REGION Network 126: DB2062.DBX17.2/3 = LT422 1P Tank Level
   // BTCS_ALARM_WORD_09_BIT_10/11                      14.13
   RUNG wire#powerrail
      "LT422 1P  TANK LEVEL ALARM"(Enable := wire#w1, Value := "20_TANKS_IP_DATA".RIO_01.SECOND_TANK.BWT_LEVEL, "Raw Value" := "IN_Level_WBT_1P", "Enable Delay Time" := "2086_Times"."Alarm Enable Delay", "High Value Release" := false, "SHORT CIRCUIT VALUE" :=, "BROKEN WIRE VALUE" :=, "VERY LOW LEVEL VALUE (LL)" :=, "LOW LEVEL VALUE (L)" := "2084_Setpoints".LT422_Lo, "HIGH LEVEL VALUE (H)" := "2084_Setpoints".LT422_Hi, "VERY HIGH LEVEL VALUE (HH)" := 32000.0, OFFSET :=, "ALARM DELAY" := "2086_Times"."LT422 Alarm Delay", "Peak Value Reset" :=, "ALARM HH" =>, "ALARM H" =>, "ALARM L" =>, "ALARM LL" =>, "ALARM READING" => %DB2062.DBX367.5, "Peak Value" =>, Alarm =>, Alarm_INT =>)   // Raw value not available for Out of Range determination
      wire#w2
      Contact( "LT422 1P  TANK LEVEL ALARM"."ALARM H" )
      Coil( %DB2062.DBX17.2 )
   END_RUNG
   RUNG wire#powerrail
      I_Contact( "2062_Warning_Data"."Water Level Override 1P" )
      { S7_Templates := "SrcType := Int" } GT_Contact(in1 := "504_Tank Grouping_DB2020"."GROUP of TANK 2", in2 := 0)
   END_RUNG wire#w1
   RUNG wire#w2
      Contact( "LT422 1P  TANK LEVEL ALARM"."ALARM L" )
      Coil( %DB2062.DBX17.3 )
   END_RUNG
   // the same network as SCL:
   "LT422 1P  TANK LEVEL ALARM"(Value := "20_TANKS_IP_DATA".RIO_01.SECOND_TANK.BWT_LEVEL,   // "502_ALM_ANALOG": Raw value not available for Out of Range determination
                           "Raw Value" := "IN_Level_WBT_1P",
                           Enable := NOT "2062_Warning_Data"."Water Level Override 1P" AND ("504_Tank Grouping_DB2020"."GROUP of TANK 2" > 0),
                           "Enable Delay Time" := "2086_Times"."Alarm Enable Delay",
                           "High Value Release" := false,
                           "LOW LEVEL VALUE (L)" := "2084_Setpoints".LT422_Lo,
                           "HIGH LEVEL VALUE (H)" := "2084_Setpoints".LT422_Hi,
                           "VERY HIGH LEVEL VALUE (HH)" := 32000.0,
                           "ALARM DELAY" := "2086_Times"."LT422 Alarm Delay",
                           "ALARM READING" => %DB2062.DBX367.5,
                           ENO => #_w1);
   %DB2062.DBX17.2 := #_w1 AND "LT422 1P  TANK LEVEL ALARM"."ALARM H";
   %DB2062.DBX17.3 := #_w1 AND "LT422 1P  TANK LEVEL ALARM"."ALARM L";
END_REGION

REGION Network 127: DB2062.DBX17.4/5 = LT421 1S Tank Level
   // BTCS_ALARM_WORD_09_BIT_12/13                                  14.14
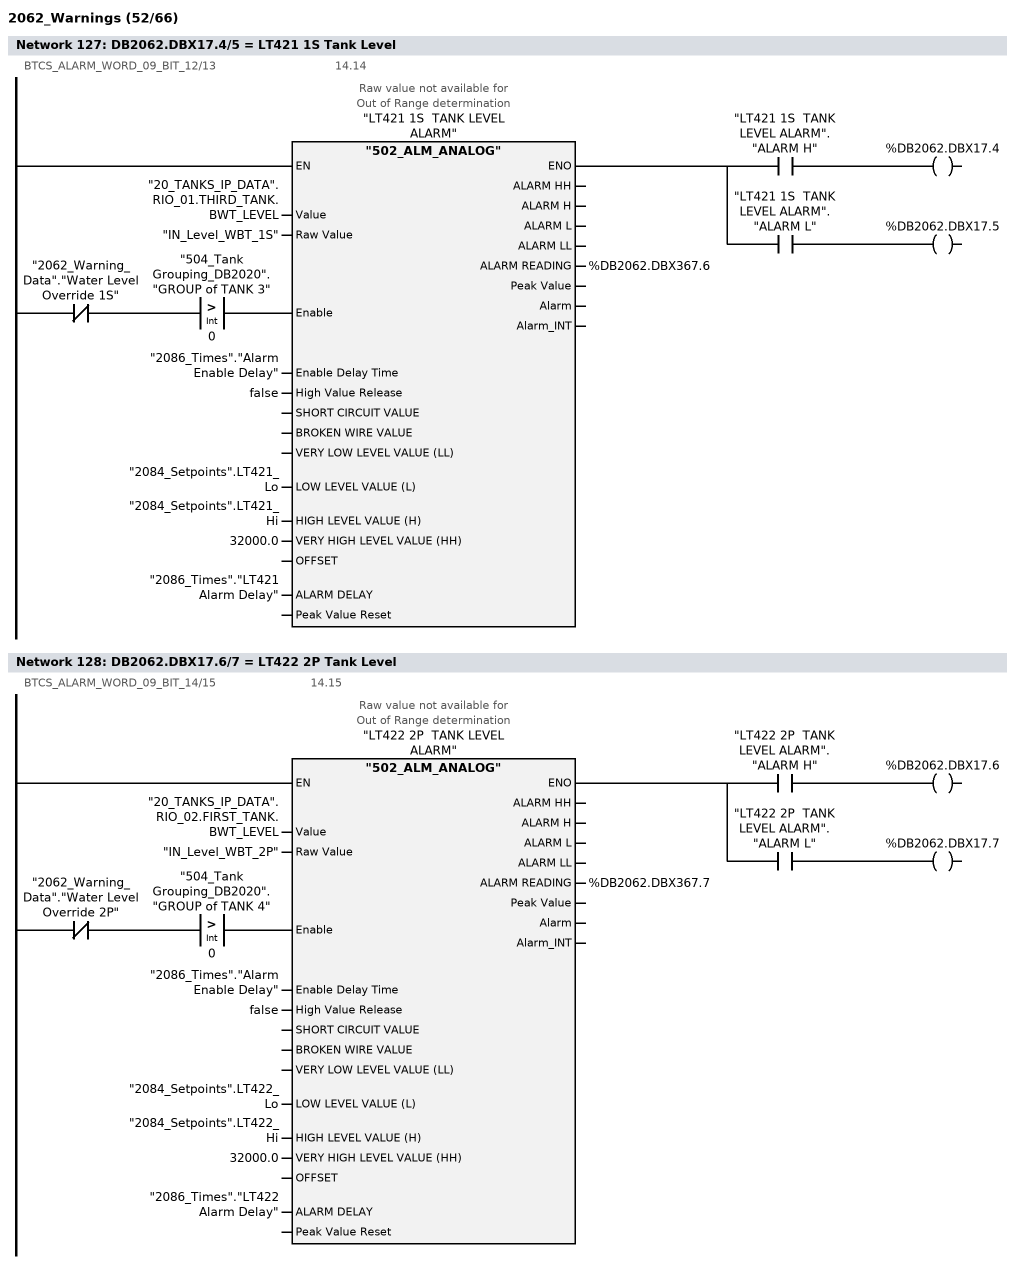
   RUNG wire#powerrail
      "LT421 1S  TANK LEVEL ALARM"(Enable := wire#w1, Value := "20_TANKS_IP_DATA".RIO_01.THIRD_TANK.BWT_LEVEL, "Raw Value" := "IN_Level_WBT_1S", "Enable Delay Time" := "2086_Times"."Alarm Enable Delay", "High Value Release" := false, "SHORT CIRCUIT VALUE" :=, "BROKEN WIRE VALUE" :=, "VERY LOW LEVEL VALUE (LL)" :=, "LOW LEVEL VALUE (L)" := "2084_Setpoints".LT421_Lo, "HIGH LEVEL VALUE (H)" := "2084_Setpoints".LT421_Hi, "VERY HIGH LEVEL VALUE (HH)" := 32000.0, OFFSET :=, "ALARM DELAY" := "2086_Times"."LT421 Alarm Delay", "Peak Value Reset" :=, "ALARM HH" =>, "ALARM H" =>, "ALARM L" =>, "ALARM LL" =>, "ALARM READING" => %DB2062.DBX367.6, "Peak Value" =>, Alarm =>, Alarm_INT =>)   // Raw value not available for Out of Range determination
      wire#w2
      Contact( "LT421 1S  TANK LEVEL ALARM"."ALARM H" )
      Coil( %DB2062.DBX17.4 )
   END_RUNG
   RUNG wire#powerrail
      I_Contact( "2062_Warning_Data"."Water Level Override 1S" )
      { S7_Templates := "SrcType := Int" } GT_Contact(in1 := "504_Tank Grouping_DB2020"."GROUP of TANK 3", in2 := 0)
   END_RUNG wire#w1
   RUNG wire#w2
      Contact( "LT421 1S  TANK LEVEL ALARM"."ALARM L" )
      Coil( %DB2062.DBX17.5 )
   END_RUNG
   // the same network as SCL:
   "LT421 1S  TANK LEVEL ALARM"(Value := "20_TANKS_IP_DATA".RIO_01.THIRD_TANK.BWT_LEVEL,   // "502_ALM_ANALOG": Raw value not available for Out of Range determination
                           "Raw Value" := "IN_Level_WBT_1S",
                           Enable := NOT "2062_Warning_Data"."Water Level Override 1S" AND ("504_Tank Grouping_DB2020"."GROUP of TANK 3" > 0),
                           "Enable Delay Time" := "2086_Times"."Alarm Enable Delay",
                           "High Value Release" := false,
                           "LOW LEVEL VALUE (L)" := "2084_Setpoints".LT421_Lo,
                           "HIGH LEVEL VALUE (H)" := "2084_Setpoints".LT421_Hi,
                           "VERY HIGH LEVEL VALUE (HH)" := 32000.0,
                           "ALARM DELAY" := "2086_Times"."LT421 Alarm Delay",
                           "ALARM READING" => %DB2062.DBX367.6,
                           ENO => #_w1);
   %DB2062.DBX17.4 := #_w1 AND "LT421 1S  TANK LEVEL ALARM"."ALARM H";
   %DB2062.DBX17.5 := #_w1 AND "LT421 1S  TANK LEVEL ALARM"."ALARM L";
END_REGION

REGION Network 128: DB2062.DBX17.6/7 = LT422 2P Tank Level
   // BTCS_ALARM_WORD_09_BIT_14/15                           14.15
   RUNG wire#powerrail
      "LT422 2P  TANK LEVEL ALARM"(Enable := wire#w1, Value := "20_TANKS_IP_DATA".RIO_02.FIRST_TANK.BWT_LEVEL, "Raw Value" := "IN_Level_WBT_2P", "Enable Delay Time" := "2086_Times"."Alarm Enable Delay", "High Value Release" := false, "SHORT CIRCUIT VALUE" :=, "BROKEN WIRE VALUE" :=, "VERY LOW LEVEL VALUE (LL)" :=, "LOW LEVEL VALUE (L)" := "2084_Setpoints".LT422_Lo, "HIGH LEVEL VALUE (H)" := "2084_Setpoints".LT422_Hi, "VERY HIGH LEVEL VALUE (HH)" := 32000.0, OFFSET :=, "ALARM DELAY" := "2086_Times"."LT422 Alarm Delay", "Peak Value Reset" :=, "ALARM HH" =>, "ALARM H" =>, "ALARM L" =>, "ALARM LL" =>, "ALARM READING" => %DB2062.DBX367.7, "Peak Value" =>, Alarm =>, Alarm_INT =>)   // Raw value not available for Out of Range determination
      wire#w2
      Contact( "LT422 2P  TANK LEVEL ALARM"."ALARM H" )
      Coil( %DB2062.DBX17.6 )
   END_RUNG
   RUNG wire#powerrail
      I_Contact( "2062_Warning_Data"."Water Level Override 2P" )
      { S7_Templates := "SrcType := Int" } GT_Contact(in1 := "504_Tank Grouping_DB2020"."GROUP of TANK 4", in2 := 0)
   END_RUNG wire#w1
   RUNG wire#w2
      Contact( "LT422 2P  TANK LEVEL ALARM"."ALARM L" )
      Coil( %DB2062.DBX17.7 )
   END_RUNG
   // the same network as SCL:
   "LT422 2P  TANK LEVEL ALARM"(Value := "20_TANKS_IP_DATA".RIO_02.FIRST_TANK.BWT_LEVEL,   // "502_ALM_ANALOG": Raw value not available for Out of Range determination
                           "Raw Value" := "IN_Level_WBT_2P",
                           Enable := NOT "2062_Warning_Data"."Water Level Override 2P" AND ("504_Tank Grouping_DB2020"."GROUP of TANK 4" > 0),
                           "Enable Delay Time" := "2086_Times"."Alarm Enable Delay",
                           "High Value Release" := false,
                           "LOW LEVEL VALUE (L)" := "2084_Setpoints".LT422_Lo,
                           "HIGH LEVEL VALUE (H)" := "2084_Setpoints".LT422_Hi,
                           "VERY HIGH LEVEL VALUE (HH)" := 32000.0,
                           "ALARM DELAY" := "2086_Times"."LT422 Alarm Delay",
                           "ALARM READING" => %DB2062.DBX367.7,
                           ENO => #_w1);
   %DB2062.DBX17.6 := #_w1 AND "LT422 2P  TANK LEVEL ALARM"."ALARM H";
   %DB2062.DBX17.7 := #_w1 AND "LT422 2P  TANK LEVEL ALARM"."ALARM L";
END_REGION

REGION Network 129: DB2062.DBX18.0/1 = LT421 2S Tank Level
   // BTCS_ALARM_WORD_10_BIT_0/1                                    15.0
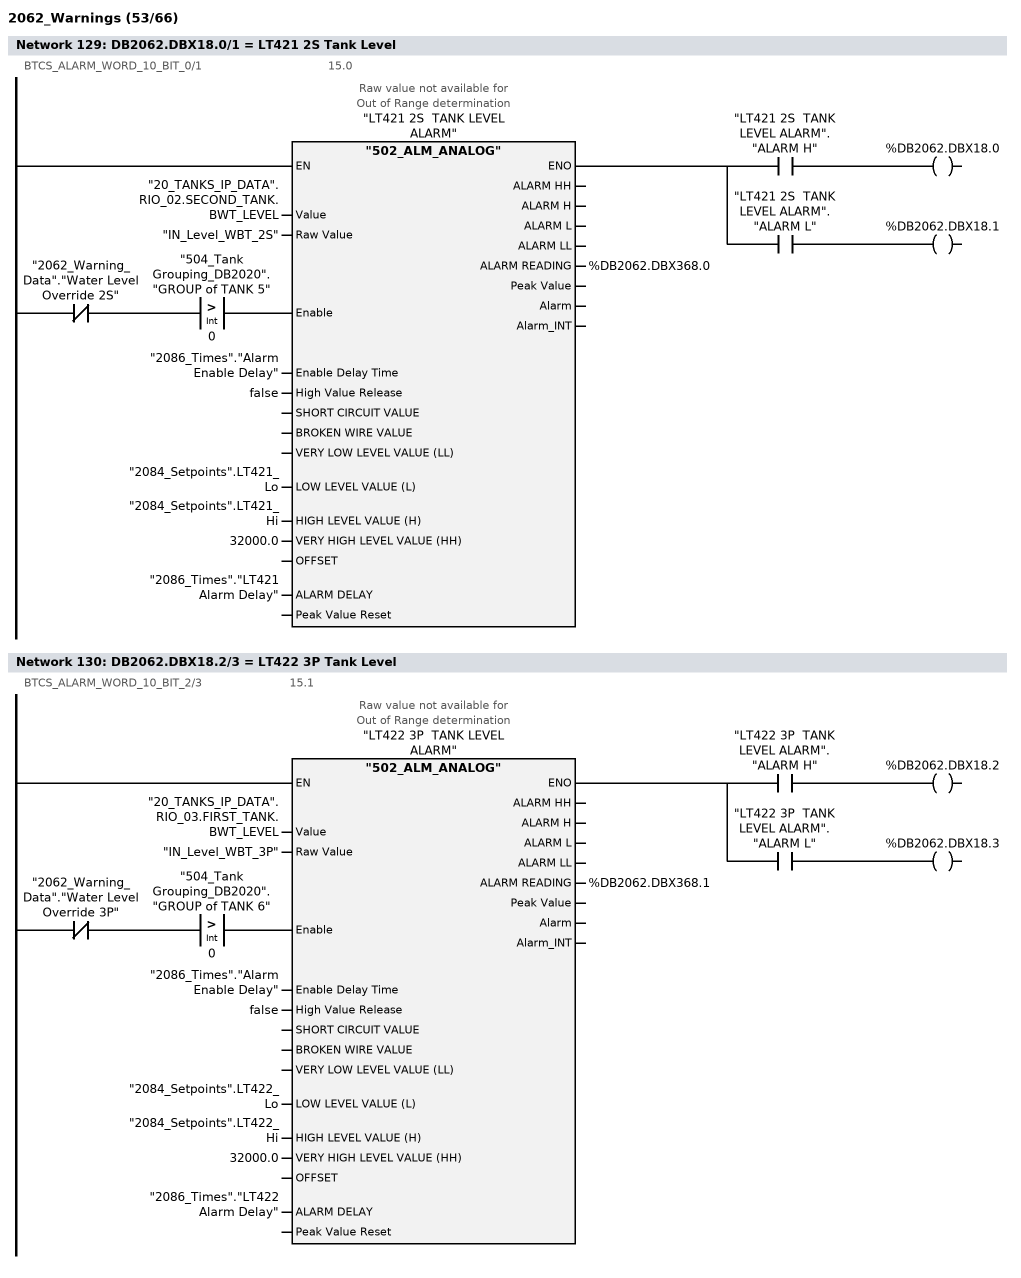
   RUNG wire#powerrail
      "LT421 2S  TANK LEVEL ALARM"(Enable := wire#w1, Value := "20_TANKS_IP_DATA".RIO_02.SECOND_TANK.BWT_LEVEL, "Raw Value" := "IN_Level_WBT_2S", "Enable Delay Time" := "2086_Times"."Alarm Enable Delay", "High Value Release" := false, "SHORT CIRCUIT VALUE" :=, "BROKEN WIRE VALUE" :=, "VERY LOW LEVEL VALUE (LL)" :=, "LOW LEVEL VALUE (L)" := "2084_Setpoints".LT421_Lo, "HIGH LEVEL VALUE (H)" := "2084_Setpoints".LT421_Hi, "VERY HIGH LEVEL VALUE (HH)" := 32000.0, OFFSET :=, "ALARM DELAY" := "2086_Times"."LT421 Alarm Delay", "Peak Value Reset" :=, "ALARM HH" =>, "ALARM H" =>, "ALARM L" =>, "ALARM LL" =>, "ALARM READING" => %DB2062.DBX368.0, "Peak Value" =>, Alarm =>, Alarm_INT =>)   // Raw value not available for Out of Range determination
      wire#w2
      Contact( "LT421 2S  TANK LEVEL ALARM"."ALARM H" )
      Coil( %DB2062.DBX18.0 )
   END_RUNG
   RUNG wire#powerrail
      I_Contact( "2062_Warning_Data"."Water Level Override 2S" )
      { S7_Templates := "SrcType := Int" } GT_Contact(in1 := "504_Tank Grouping_DB2020"."GROUP of TANK 5", in2 := 0)
   END_RUNG wire#w1
   RUNG wire#w2
      Contact( "LT421 2S  TANK LEVEL ALARM"."ALARM L" )
      Coil( %DB2062.DBX18.1 )
   END_RUNG
   // the same network as SCL:
   "LT421 2S  TANK LEVEL ALARM"(Value := "20_TANKS_IP_DATA".RIO_02.SECOND_TANK.BWT_LEVEL,   // "502_ALM_ANALOG": Raw value not available for Out of Range determination
                           "Raw Value" := "IN_Level_WBT_2S",
                           Enable := NOT "2062_Warning_Data"."Water Level Override 2S" AND ("504_Tank Grouping_DB2020"."GROUP of TANK 5" > 0),
                           "Enable Delay Time" := "2086_Times"."Alarm Enable Delay",
                           "High Value Release" := false,
                           "LOW LEVEL VALUE (L)" := "2084_Setpoints".LT421_Lo,
                           "HIGH LEVEL VALUE (H)" := "2084_Setpoints".LT421_Hi,
                           "VERY HIGH LEVEL VALUE (HH)" := 32000.0,
                           "ALARM DELAY" := "2086_Times"."LT421 Alarm Delay",
                           "ALARM READING" => %DB2062.DBX368.0,
                           ENO => #_w1);
   %DB2062.DBX18.0 := #_w1 AND "LT421 2S  TANK LEVEL ALARM"."ALARM H";
   %DB2062.DBX18.1 := #_w1 AND "LT421 2S  TANK LEVEL ALARM"."ALARM L";
END_REGION

REGION Network 130: DB2062.DBX18.2/3 = LT422 3P Tank Level
   // BTCS_ALARM_WORD_10_BIT_2/3                         15.1
   RUNG wire#powerrail
      "LT422 3P  TANK LEVEL ALARM"(Enable := wire#w1, Value := "20_TANKS_IP_DATA".RIO_03.FIRST_TANK.BWT_LEVEL, "Raw Value" := "IN_Level_WBT_3P", "Enable Delay Time" := "2086_Times"."Alarm Enable Delay", "High Value Release" := false, "SHORT CIRCUIT VALUE" :=, "BROKEN WIRE VALUE" :=, "VERY LOW LEVEL VALUE (LL)" :=, "LOW LEVEL VALUE (L)" := "2084_Setpoints".LT422_Lo, "HIGH LEVEL VALUE (H)" := "2084_Setpoints".LT422_Hi, "VERY HIGH LEVEL VALUE (HH)" := 32000.0, OFFSET :=, "ALARM DELAY" := "2086_Times"."LT422 Alarm Delay", "Peak Value Reset" :=, "ALARM HH" =>, "ALARM H" =>, "ALARM L" =>, "ALARM LL" =>, "ALARM READING" => %DB2062.DBX368.1, "Peak Value" =>, Alarm =>, Alarm_INT =>)   // Raw value not available for Out of Range determination
      wire#w2
      Contact( "LT422 3P  TANK LEVEL ALARM"."ALARM H" )
      Coil( %DB2062.DBX18.2 )
   END_RUNG
   RUNG wire#powerrail
      I_Contact( "2062_Warning_Data"."Water Level Override 3P" )
      { S7_Templates := "SrcType := Int" } GT_Contact(in1 := "504_Tank Grouping_DB2020"."GROUP of TANK 6", in2 := 0)
   END_RUNG wire#w1
   RUNG wire#w2
      Contact( "LT422 3P  TANK LEVEL ALARM"."ALARM L" )
      Coil( %DB2062.DBX18.3 )
   END_RUNG
   // the same network as SCL:
   "LT422 3P  TANK LEVEL ALARM"(Value := "20_TANKS_IP_DATA".RIO_03.FIRST_TANK.BWT_LEVEL,   // "502_ALM_ANALOG": Raw value not available for Out of Range determination
                           "Raw Value" := "IN_Level_WBT_3P",
                           Enable := NOT "2062_Warning_Data"."Water Level Override 3P" AND ("504_Tank Grouping_DB2020"."GROUP of TANK 6" > 0),
                           "Enable Delay Time" := "2086_Times"."Alarm Enable Delay",
                           "High Value Release" := false,
                           "LOW LEVEL VALUE (L)" := "2084_Setpoints".LT422_Lo,
                           "HIGH LEVEL VALUE (H)" := "2084_Setpoints".LT422_Hi,
                           "VERY HIGH LEVEL VALUE (HH)" := 32000.0,
                           "ALARM DELAY" := "2086_Times"."LT422 Alarm Delay",
                           "ALARM READING" => %DB2062.DBX368.1,
                           ENO => #_w1);
   %DB2062.DBX18.2 := #_w1 AND "LT422 3P  TANK LEVEL ALARM"."ALARM H";
   %DB2062.DBX18.3 := #_w1 AND "LT422 3P  TANK LEVEL ALARM"."ALARM L";
END_REGION

REGION Network 131: DB2062.DBX18.4/5 = LT421 3S Tank Level
   // BTCS_ALARM_WORD_10_BIT_4/5                               15.2
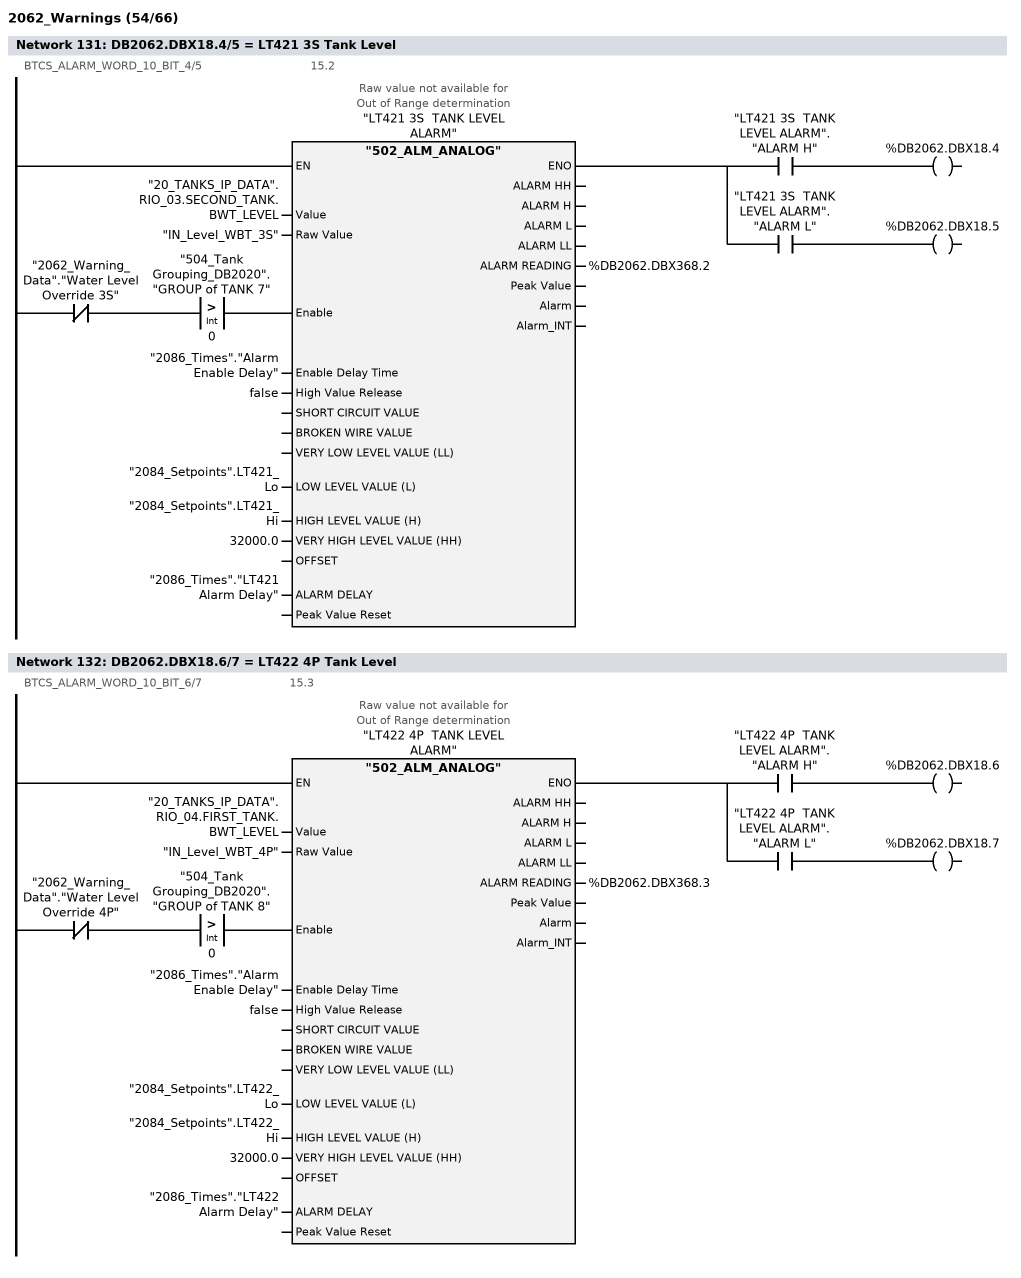
   RUNG wire#powerrail
      "LT421 3S  TANK LEVEL ALARM"(Enable := wire#w1, Value := "20_TANKS_IP_DATA".RIO_03.SECOND_TANK.BWT_LEVEL, "Raw Value" := "IN_Level_WBT_3S", "Enable Delay Time" := "2086_Times"."Alarm Enable Delay", "High Value Release" := false, "SHORT CIRCUIT VALUE" :=, "BROKEN WIRE VALUE" :=, "VERY LOW LEVEL VALUE (LL)" :=, "LOW LEVEL VALUE (L)" := "2084_Setpoints".LT421_Lo, "HIGH LEVEL VALUE (H)" := "2084_Setpoints".LT421_Hi, "VERY HIGH LEVEL VALUE (HH)" := 32000.0, OFFSET :=, "ALARM DELAY" := "2086_Times"."LT421 Alarm Delay", "Peak Value Reset" :=, "ALARM HH" =>, "ALARM H" =>, "ALARM L" =>, "ALARM LL" =>, "ALARM READING" => %DB2062.DBX368.2, "Peak Value" =>, Alarm =>, Alarm_INT =>)   // Raw value not available for Out of Range determination
      wire#w2
      Contact( "LT421 3S  TANK LEVEL ALARM"."ALARM H" )
      Coil( %DB2062.DBX18.4 )
   END_RUNG
   RUNG wire#powerrail
      I_Contact( "2062_Warning_Data"."Water Level Override 3S" )
      { S7_Templates := "SrcType := Int" } GT_Contact(in1 := "504_Tank Grouping_DB2020"."GROUP of TANK 7", in2 := 0)
   END_RUNG wire#w1
   RUNG wire#w2
      Contact( "LT421 3S  TANK LEVEL ALARM"."ALARM L" )
      Coil( %DB2062.DBX18.5 )
   END_RUNG
   // the same network as SCL:
   "LT421 3S  TANK LEVEL ALARM"(Value := "20_TANKS_IP_DATA".RIO_03.SECOND_TANK.BWT_LEVEL,   // "502_ALM_ANALOG": Raw value not available for Out of Range determination
                           "Raw Value" := "IN_Level_WBT_3S",
                           Enable := NOT "2062_Warning_Data"."Water Level Override 3S" AND ("504_Tank Grouping_DB2020"."GROUP of TANK 7" > 0),
                           "Enable Delay Time" := "2086_Times"."Alarm Enable Delay",
                           "High Value Release" := false,
                           "LOW LEVEL VALUE (L)" := "2084_Setpoints".LT421_Lo,
                           "HIGH LEVEL VALUE (H)" := "2084_Setpoints".LT421_Hi,
                           "VERY HIGH LEVEL VALUE (HH)" := 32000.0,
                           "ALARM DELAY" := "2086_Times"."LT421 Alarm Delay",
                           "ALARM READING" => %DB2062.DBX368.2,
                           ENO => #_w1);
   %DB2062.DBX18.4 := #_w1 AND "LT421 3S  TANK LEVEL ALARM"."ALARM H";
   %DB2062.DBX18.5 := #_w1 AND "LT421 3S  TANK LEVEL ALARM"."ALARM L";
END_REGION

REGION Network 132: DB2062.DBX18.6/7 = LT422 4P Tank Level
   // BTCS_ALARM_WORD_10_BIT_6/7                         15.3
   RUNG wire#powerrail
      "LT422 4P  TANK LEVEL ALARM"(Enable := wire#w1, Value := "20_TANKS_IP_DATA".RIO_04.FIRST_TANK.BWT_LEVEL, "Raw Value" := "IN_Level_WBT_4P", "Enable Delay Time" := "2086_Times"."Alarm Enable Delay", "High Value Release" := false, "SHORT CIRCUIT VALUE" :=, "BROKEN WIRE VALUE" :=, "VERY LOW LEVEL VALUE (LL)" :=, "LOW LEVEL VALUE (L)" := "2084_Setpoints".LT422_Lo, "HIGH LEVEL VALUE (H)" := "2084_Setpoints".LT422_Hi, "VERY HIGH LEVEL VALUE (HH)" := 32000.0, OFFSET :=, "ALARM DELAY" := "2086_Times"."LT422 Alarm Delay", "Peak Value Reset" :=, "ALARM HH" =>, "ALARM H" =>, "ALARM L" =>, "ALARM LL" =>, "ALARM READING" => %DB2062.DBX368.3, "Peak Value" =>, Alarm =>, Alarm_INT =>)   // Raw value not available for Out of Range determination
      wire#w2
      Contact( "LT422 4P  TANK LEVEL ALARM"."ALARM H" )
      Coil( %DB2062.DBX18.6 )
   END_RUNG
   RUNG wire#powerrail
      I_Contact( "2062_Warning_Data"."Water Level Override 4P" )
      { S7_Templates := "SrcType := Int" } GT_Contact(in1 := "504_Tank Grouping_DB2020"."GROUP of TANK 8", in2 := 0)
   END_RUNG wire#w1
   RUNG wire#w2
      Contact( "LT422 4P  TANK LEVEL ALARM"."ALARM L" )
      Coil( %DB2062.DBX18.7 )
   END_RUNG
   // the same network as SCL:
   "LT422 4P  TANK LEVEL ALARM"(Value := "20_TANKS_IP_DATA".RIO_04.FIRST_TANK.BWT_LEVEL,   // "502_ALM_ANALOG": Raw value not available for Out of Range determination
                           "Raw Value" := "IN_Level_WBT_4P",
                           Enable := NOT "2062_Warning_Data"."Water Level Override 4P" AND ("504_Tank Grouping_DB2020"."GROUP of TANK 8" > 0),
                           "Enable Delay Time" := "2086_Times"."Alarm Enable Delay",
                           "High Value Release" := false,
                           "LOW LEVEL VALUE (L)" := "2084_Setpoints".LT422_Lo,
                           "HIGH LEVEL VALUE (H)" := "2084_Setpoints".LT422_Hi,
                           "VERY HIGH LEVEL VALUE (HH)" := 32000.0,
                           "ALARM DELAY" := "2086_Times"."LT422 Alarm Delay",
                           "ALARM READING" => %DB2062.DBX368.3,
                           ENO => #_w1);
   %DB2062.DBX18.6 := #_w1 AND "LT422 4P  TANK LEVEL ALARM"."ALARM H";
   %DB2062.DBX18.7 := #_w1 AND "LT422 4P  TANK LEVEL ALARM"."ALARM L";
END_REGION

REGION Network 133: DB2062.DBX19.0/1 = LT421 4S Tank Level
   // BTCS_ALARM_WORD_10_BIT_8/9                     15.4
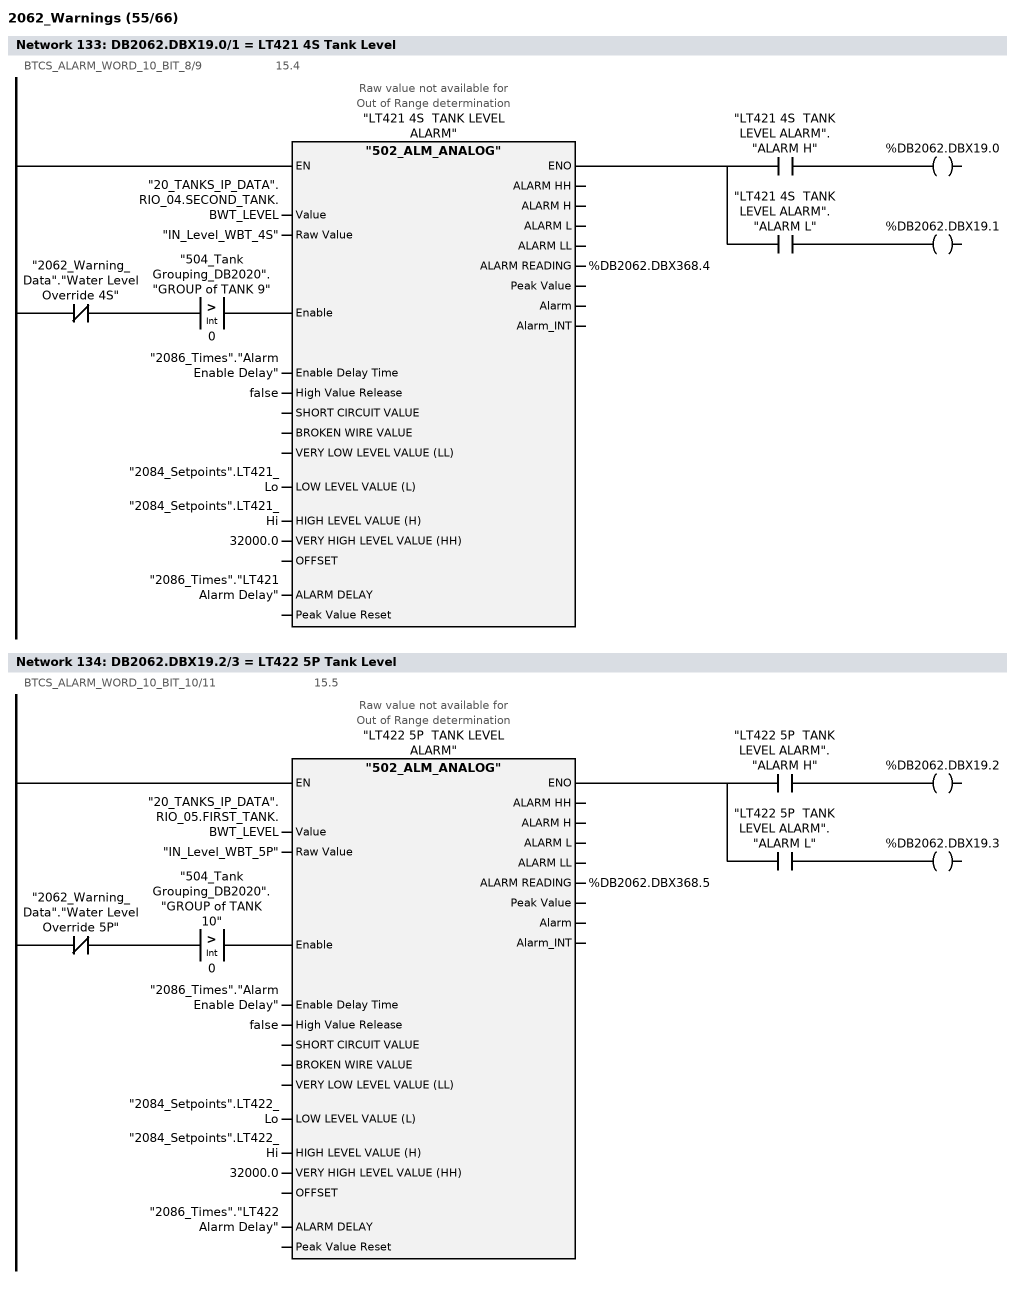
   RUNG wire#powerrail
      "LT421 4S  TANK LEVEL ALARM"(Enable := wire#w1, Value := "20_TANKS_IP_DATA".RIO_04.SECOND_TANK.BWT_LEVEL, "Raw Value" := "IN_Level_WBT_4S", "Enable Delay Time" := "2086_Times"."Alarm Enable Delay", "High Value Release" := false, "SHORT CIRCUIT VALUE" :=, "BROKEN WIRE VALUE" :=, "VERY LOW LEVEL VALUE (LL)" :=, "LOW LEVEL VALUE (L)" := "2084_Setpoints".LT421_Lo, "HIGH LEVEL VALUE (H)" := "2084_Setpoints".LT421_Hi, "VERY HIGH LEVEL VALUE (HH)" := 32000.0, OFFSET :=, "ALARM DELAY" := "2086_Times"."LT421 Alarm Delay", "Peak Value Reset" :=, "ALARM HH" =>, "ALARM H" =>, "ALARM L" =>, "ALARM LL" =>, "ALARM READING" => %DB2062.DBX368.4, "Peak Value" =>, Alarm =>, Alarm_INT =>)   // Raw value not available for Out of Range determination
      wire#w2
      Contact( "LT421 4S  TANK LEVEL ALARM"."ALARM H" )
      Coil( %DB2062.DBX19.0 )
   END_RUNG
   RUNG wire#powerrail
      I_Contact( "2062_Warning_Data"."Water Level Override 4S" )
      { S7_Templates := "SrcType := Int" } GT_Contact(in1 := "504_Tank Grouping_DB2020"."GROUP of TANK 9", in2 := 0)
   END_RUNG wire#w1
   RUNG wire#w2
      Contact( "LT421 4S  TANK LEVEL ALARM"."ALARM L" )
      Coil( %DB2062.DBX19.1 )
   END_RUNG
   // the same network as SCL:
   "LT421 4S  TANK LEVEL ALARM"(Value := "20_TANKS_IP_DATA".RIO_04.SECOND_TANK.BWT_LEVEL,   // "502_ALM_ANALOG": Raw value not available for Out of Range determination
                           "Raw Value" := "IN_Level_WBT_4S",
                           Enable := NOT "2062_Warning_Data"."Water Level Override 4S" AND ("504_Tank Grouping_DB2020"."GROUP of TANK 9" > 0),
                           "Enable Delay Time" := "2086_Times"."Alarm Enable Delay",
                           "High Value Release" := false,
                           "LOW LEVEL VALUE (L)" := "2084_Setpoints".LT421_Lo,
                           "HIGH LEVEL VALUE (H)" := "2084_Setpoints".LT421_Hi,
                           "VERY HIGH LEVEL VALUE (HH)" := 32000.0,
                           "ALARM DELAY" := "2086_Times"."LT421 Alarm Delay",
                           "ALARM READING" => %DB2062.DBX368.4,
                           ENO => #_w1);
   %DB2062.DBX19.0 := #_w1 AND "LT421 4S  TANK LEVEL ALARM"."ALARM H";
   %DB2062.DBX19.1 := #_w1 AND "LT421 4S  TANK LEVEL ALARM"."ALARM L";
END_REGION

REGION Network 134: DB2062.DBX19.2/3 = LT422 5P Tank Level
   // BTCS_ALARM_WORD_10_BIT_10/11                            15.5
   RUNG wire#powerrail
      "LT422 5P  TANK LEVEL ALARM"(Enable := wire#w1, Value := "20_TANKS_IP_DATA".RIO_05.FIRST_TANK.BWT_LEVEL, "Raw Value" := "IN_Level_WBT_5P", "Enable Delay Time" := "2086_Times"."Alarm Enable Delay", "High Value Release" := false, "SHORT CIRCUIT VALUE" :=, "BROKEN WIRE VALUE" :=, "VERY LOW LEVEL VALUE (LL)" :=, "LOW LEVEL VALUE (L)" := "2084_Setpoints".LT422_Lo, "HIGH LEVEL VALUE (H)" := "2084_Setpoints".LT422_Hi, "VERY HIGH LEVEL VALUE (HH)" := 32000.0, OFFSET :=, "ALARM DELAY" := "2086_Times"."LT422 Alarm Delay", "Peak Value Reset" :=, "ALARM HH" =>, "ALARM H" =>, "ALARM L" =>, "ALARM LL" =>, "ALARM READING" => %DB2062.DBX368.5, "Peak Value" =>, Alarm =>, Alarm_INT =>)   // Raw value not available for Out of Range determination
      wire#w2
      Contact( "LT422 5P  TANK LEVEL ALARM"."ALARM H" )
      Coil( %DB2062.DBX19.2 )
   END_RUNG
   RUNG wire#powerrail
      I_Contact( "2062_Warning_Data"."Water Level Override 5P" )
      { S7_Templates := "SrcType := Int" } GT_Contact(in1 := "504_Tank Grouping_DB2020"."GROUP of TANK 10", in2 := 0)
   END_RUNG wire#w1
   RUNG wire#w2
      Contact( "LT422 5P  TANK LEVEL ALARM"."ALARM L" )
      Coil( %DB2062.DBX19.3 )
   END_RUNG
   // the same network as SCL:
   "LT422 5P  TANK LEVEL ALARM"(Value := "20_TANKS_IP_DATA".RIO_05.FIRST_TANK.BWT_LEVEL,   // "502_ALM_ANALOG": Raw value not available for Out of Range determination
                           "Raw Value" := "IN_Level_WBT_5P",
                           Enable := NOT "2062_Warning_Data"."Water Level Override 5P" AND ("504_Tank Grouping_DB2020"."GROUP of TANK 10" > 0),
                           "Enable Delay Time" := "2086_Times"."Alarm Enable Delay",
                           "High Value Release" := false,
                           "LOW LEVEL VALUE (L)" := "2084_Setpoints".LT422_Lo,
                           "HIGH LEVEL VALUE (H)" := "2084_Setpoints".LT422_Hi,
                           "VERY HIGH LEVEL VALUE (HH)" := 32000.0,
                           "ALARM DELAY" := "2086_Times"."LT422 Alarm Delay",
                           "ALARM READING" => %DB2062.DBX368.5,
                           ENO => #_w1);
   %DB2062.DBX19.2 := #_w1 AND "LT422 5P  TANK LEVEL ALARM"."ALARM H";
   %DB2062.DBX19.3 := #_w1 AND "LT422 5P  TANK LEVEL ALARM"."ALARM L";
END_REGION

REGION Network 135: DB2062.DBX19.4/5 = LT421 5S Tank Level
   // BTCS_ALARM_WORD_10_BIT_12/13                          15.6
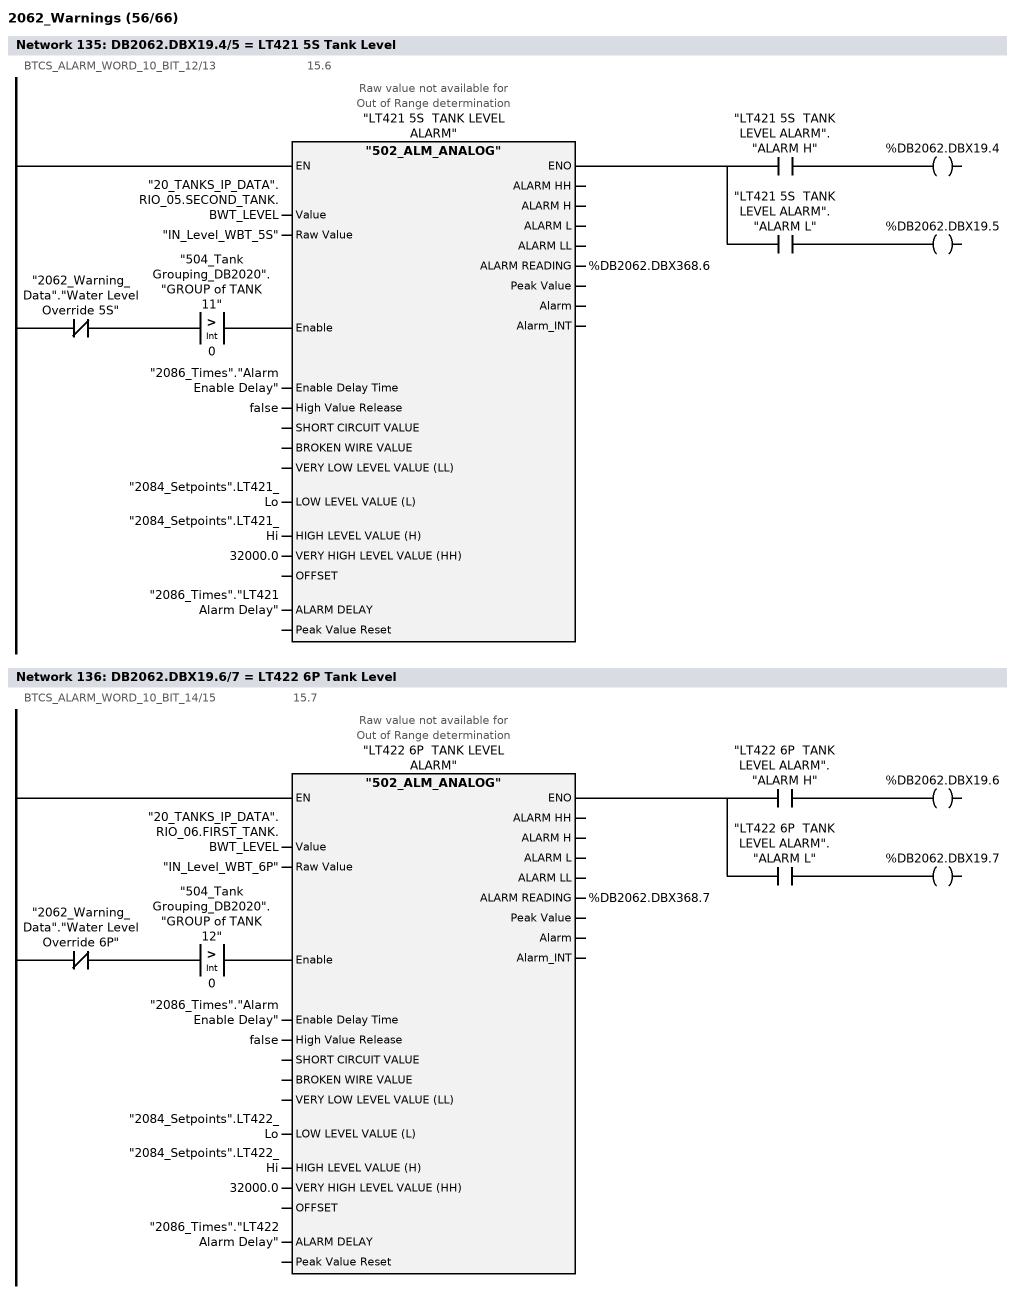
   RUNG wire#powerrail
      "LT421 5S  TANK LEVEL ALARM"(Enable := wire#w1, Value := "20_TANKS_IP_DATA".RIO_05.SECOND_TANK.BWT_LEVEL, "Raw Value" := "IN_Level_WBT_5S", "Enable Delay Time" := "2086_Times"."Alarm Enable Delay", "High Value Release" := false, "SHORT CIRCUIT VALUE" :=, "BROKEN WIRE VALUE" :=, "VERY LOW LEVEL VALUE (LL)" :=, "LOW LEVEL VALUE (L)" := "2084_Setpoints".LT421_Lo, "HIGH LEVEL VALUE (H)" := "2084_Setpoints".LT421_Hi, "VERY HIGH LEVEL VALUE (HH)" := 32000.0, OFFSET :=, "ALARM DELAY" := "2086_Times"."LT421 Alarm Delay", "Peak Value Reset" :=, "ALARM HH" =>, "ALARM H" =>, "ALARM L" =>, "ALARM LL" =>, "ALARM READING" => %DB2062.DBX368.6, "Peak Value" =>, Alarm =>, Alarm_INT =>)   // Raw value not available for Out of Range determination
      wire#w2
      Contact( "LT421 5S  TANK LEVEL ALARM"."ALARM H" )
      Coil( %DB2062.DBX19.4 )
   END_RUNG
   RUNG wire#powerrail
      I_Contact( "2062_Warning_Data"."Water Level Override 5S" )
      { S7_Templates := "SrcType := Int" } GT_Contact(in1 := "504_Tank Grouping_DB2020"."GROUP of TANK 11", in2 := 0)
   END_RUNG wire#w1
   RUNG wire#w2
      Contact( "LT421 5S  TANK LEVEL ALARM"."ALARM L" )
      Coil( %DB2062.DBX19.5 )
   END_RUNG
   // the same network as SCL:
   "LT421 5S  TANK LEVEL ALARM"(Value := "20_TANKS_IP_DATA".RIO_05.SECOND_TANK.BWT_LEVEL,   // "502_ALM_ANALOG": Raw value not available for Out of Range determination
                           "Raw Value" := "IN_Level_WBT_5S",
                           Enable := NOT "2062_Warning_Data"."Water Level Override 5S" AND ("504_Tank Grouping_DB2020"."GROUP of TANK 11" > 0),
                           "Enable Delay Time" := "2086_Times"."Alarm Enable Delay",
                           "High Value Release" := false,
                           "LOW LEVEL VALUE (L)" := "2084_Setpoints".LT421_Lo,
                           "HIGH LEVEL VALUE (H)" := "2084_Setpoints".LT421_Hi,
                           "VERY HIGH LEVEL VALUE (HH)" := 32000.0,
                           "ALARM DELAY" := "2086_Times"."LT421 Alarm Delay",
                           "ALARM READING" => %DB2062.DBX368.6,
                           ENO => #_w1);
   %DB2062.DBX19.4 := #_w1 AND "LT421 5S  TANK LEVEL ALARM"."ALARM H";
   %DB2062.DBX19.5 := #_w1 AND "LT421 5S  TANK LEVEL ALARM"."ALARM L";
END_REGION

REGION Network 136: DB2062.DBX19.6/7 = LT422 6P Tank Level
   // BTCS_ALARM_WORD_10_BIT_14/15                      15.7
   RUNG wire#powerrail
      "LT422 6P  TANK LEVEL ALARM"(Enable := wire#w1, Value := "20_TANKS_IP_DATA".RIO_06.FIRST_TANK.BWT_LEVEL, "Raw Value" := "IN_Level_WBT_6P", "Enable Delay Time" := "2086_Times"."Alarm Enable Delay", "High Value Release" := false, "SHORT CIRCUIT VALUE" :=, "BROKEN WIRE VALUE" :=, "VERY LOW LEVEL VALUE (LL)" :=, "LOW LEVEL VALUE (L)" := "2084_Setpoints".LT422_Lo, "HIGH LEVEL VALUE (H)" := "2084_Setpoints".LT422_Hi, "VERY HIGH LEVEL VALUE (HH)" := 32000.0, OFFSET :=, "ALARM DELAY" := "2086_Times"."LT422 Alarm Delay", "Peak Value Reset" :=, "ALARM HH" =>, "ALARM H" =>, "ALARM L" =>, "ALARM LL" =>, "ALARM READING" => %DB2062.DBX368.7, "Peak Value" =>, Alarm =>, Alarm_INT =>)   // Raw value not available for Out of Range determination
      wire#w2
      Contact( "LT422 6P  TANK LEVEL ALARM"."ALARM H" )
      Coil( %DB2062.DBX19.6 )
   END_RUNG
   RUNG wire#powerrail
      I_Contact( "2062_Warning_Data"."Water Level Override 6P" )
      { S7_Templates := "SrcType := Int" } GT_Contact(in1 := "504_Tank Grouping_DB2020"."GROUP of TANK 12", in2 := 0)
   END_RUNG wire#w1
   RUNG wire#w2
      Contact( "LT422 6P  TANK LEVEL ALARM"."ALARM L" )
      Coil( %DB2062.DBX19.7 )
   END_RUNG
   // the same network as SCL:
   "LT422 6P  TANK LEVEL ALARM"(Value := "20_TANKS_IP_DATA".RIO_06.FIRST_TANK.BWT_LEVEL,   // "502_ALM_ANALOG": Raw value not available for Out of Range determination
                           "Raw Value" := "IN_Level_WBT_6P",
                           Enable := NOT "2062_Warning_Data"."Water Level Override 6P" AND ("504_Tank Grouping_DB2020"."GROUP of TANK 12" > 0),
                           "Enable Delay Time" := "2086_Times"."Alarm Enable Delay",
                           "High Value Release" := false,
                           "LOW LEVEL VALUE (L)" := "2084_Setpoints".LT422_Lo,
                           "HIGH LEVEL VALUE (H)" := "2084_Setpoints".LT422_Hi,
                           "VERY HIGH LEVEL VALUE (HH)" := 32000.0,
                           "ALARM DELAY" := "2086_Times"."LT422 Alarm Delay",
                           "ALARM READING" => %DB2062.DBX368.7,
                           ENO => #_w1);
   %DB2062.DBX19.6 := #_w1 AND "LT422 6P  TANK LEVEL ALARM"."ALARM H";
   %DB2062.DBX19.7 := #_w1 AND "LT422 6P  TANK LEVEL ALARM"."ALARM L";
END_REGION

REGION Network 137: DB2062.DBX20.0/1 = LT421 6S Tank Level
   // BTCS_ALARM_WORD_11_BIT_0/1                  15.8